(* Logix 5000 project; controller FV vendor 1 type 14 code 217 rev 31.11; software revision 31.00; part 32 of 63 *)
(* tags used below, declared in another part *)
   CWD : CHECKWORD_FLAGS;
   FR_data_file_value_to_move : DINT;
   FR_DEFOAM : PlantItem;   // DEFOAM
   FR_N120 : INT[265];   // YEAST CROP Yeast Cropping Main
   FR_N120_17_0_Storagebit : BOOL;
   FR_N120_17_1_Storagebit : BOOL;
   FR_N120_17_2_Storagebit : BOOL;
   FR_N120_17_3_Storagebit : BOOL;
   FR_N120_17_4_Storagebit : BOOL;
   FR_N120_17_5_Storagebit : BOOL;
   FR_N14 : INT[265];   // MVFV CIP Comms to MVFV CIP Un it PLC
   FR_N140 : INT[265];   // CIP
   FR_N150 : INT[265];   // Original N File From SLC, No Description Available
   FR_N20 : INT[265];   // GENERAL General Purpose Setp oints
   FR_N210 : INT[265];   // ANALOG_OUT Analog Outputs
   FR_N255 : INT[265];   // CHECKWORDS
   FR_N99 : INT[265];   // COMMENT Comment Lines
   FR_SFile : INT[255];   // SLC Equivalent System File, So Original Code Can Remain
   FR_T121 : TIMER[255];   // YEAST CROP
   FR_T144 : TIMER[255];   // CIP
   FR_T4 : TIMER[255];   // TIMER
   FR_VB1_AV02 : PlantItem;   // VB1_AV02
   FR_VB1_AV04 : PlantItem;   // VB1_AV04
   FR_VB1_AV07 : PlantItem;   // VB1_AV07
   FR_VB2_AV03 : PlantItem;   // VB2_AV03
   FR_VB3_AV03 : PlantItem;   // VB3_AV03
   FR_YC_1 : PlantItem;   // YC_1
   FR_YC_2 : PlantItem;   // YC_2
   FR_YC_IN2 : PlantItem;   // YC_IN2
   FR_YC_LL : PlantItem;   // YC_LL
   FR_YEAST_121_TEMPREAL : REAL;
   FR_YM_P01 : PlantItem;   // YM_P01
   FR_YM_P02 : PlantItem;   // YM_P02
   FR_YM_P03 : PlantItem;   // YM_P03
   FR_YP1_CIP : PlantItem;   // YP1_CIP
   FR_YP2_CIP : PlantItem;   // YP2_CIP
   FR_YP3_CIP : PlantItem;   // YP3_CIP
   scale_analog_result : REAL;
   Test_Cropping_done : BOOL;
(* FR_Common, continued *)

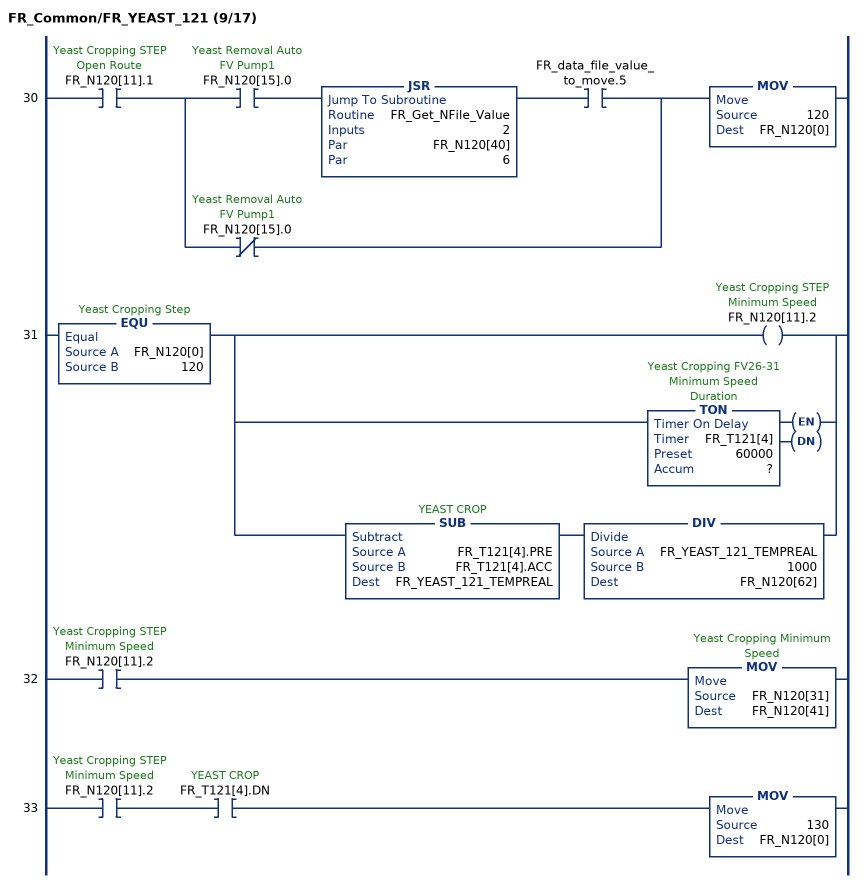
   30: XIC(FR_N120[11].1)[XIC(FR_N120[15].0) JSR(FR_Get_NFile_Value,2,FR_N120[40],6) XIC(FR_data_file_value_to_move.5) ,XIO(FR_N120[15].0) ]MOV(120,FR_N120[0]);
   31: EQU(FR_N120[0],120)[OTE(FR_N120[11].2) ,TON(FR_T121[4],?,?) ,SUB(FR_T121[4].PRE,FR_T121[4].ACC,FR_YEAST_121_TEMPREAL) DIV(FR_YEAST_121_TEMPREAL,1000,FR_N120[62]) ];
   32: XIC(FR_N120[11].2)MOV(FR_N120[31],FR_N120[41]);
   33: XIC(FR_N120[11].2)XIC(FR_T121[4].DN)MOV(130,FR_N120[0]);
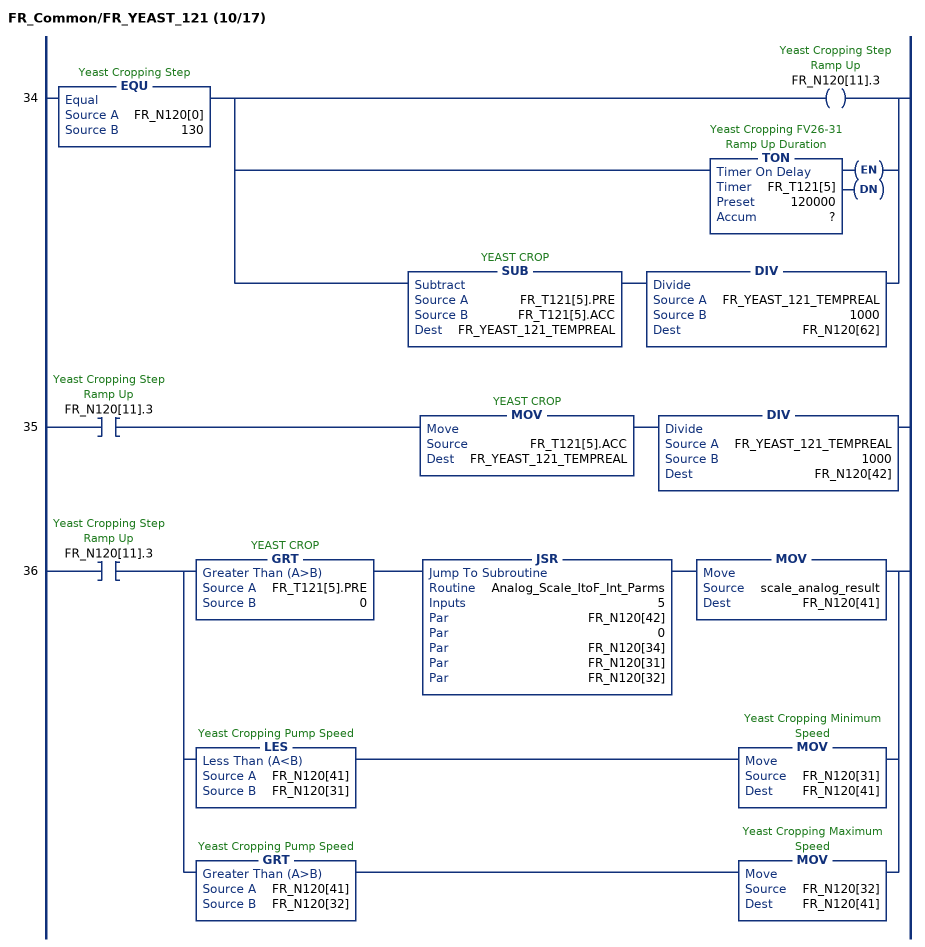
   34: EQU(FR_N120[0],130)[OTE(FR_N120[11].3) ,TON(FR_T121[5],?,?) ,SUB(FR_T121[5].PRE,FR_T121[5].ACC,FR_YEAST_121_TEMPREAL) DIV(FR_YEAST_121_TEMPREAL,1000,FR_N120[62]) ];
   35: XIC(FR_N120[11].3)MOV(FR_T121[5].ACC,FR_YEAST_121_TEMPREAL)DIV(FR_YEAST_121_TEMPREAL,1000,FR_N120[42]);
   36: XIC(FR_N120[11].3)[GRT(FR_T121[5].PRE,0) JSR(Analog_Scale_ItoF_Int_Parms,5,FR_N120[42],0,FR_N120[34],FR_N120[31],FR_N120[32]) MOV(scale_analog_result,FR_N120[41]) ,LES(FR_N120[41],FR_N120[31]) MOV(FR_N120[31],FR_N120[41]) ,GRT(FR_N120[41],FR_N120[32]) MOV(FR_N120[32],FR_N120[41]) ];
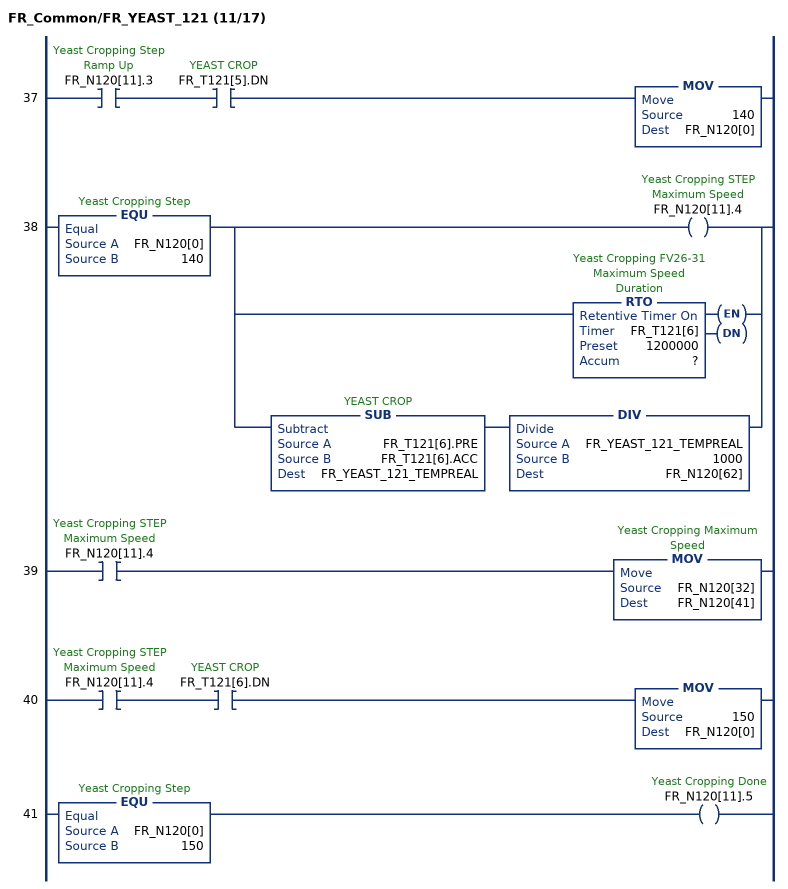
   37: XIC(FR_N120[11].3)XIC(FR_T121[5].DN)MOV(140,FR_N120[0]);
   38: EQU(FR_N120[0],140)[OTE(FR_N120[11].4) ,RTO(FR_T121[6],?,?) ,SUB(FR_T121[6].PRE,FR_T121[6].ACC,FR_YEAST_121_TEMPREAL) DIV(FR_YEAST_121_TEMPREAL,1000,FR_N120[62]) ];
   39: XIC(FR_N120[11].4)MOV(FR_N120[32],FR_N120[41]);
   40: XIC(FR_N120[11].4)XIC(FR_T121[6].DN)MOV(150,FR_N120[0]);
   41: EQU(FR_N120[0],150)OTE(FR_N120[11].5);
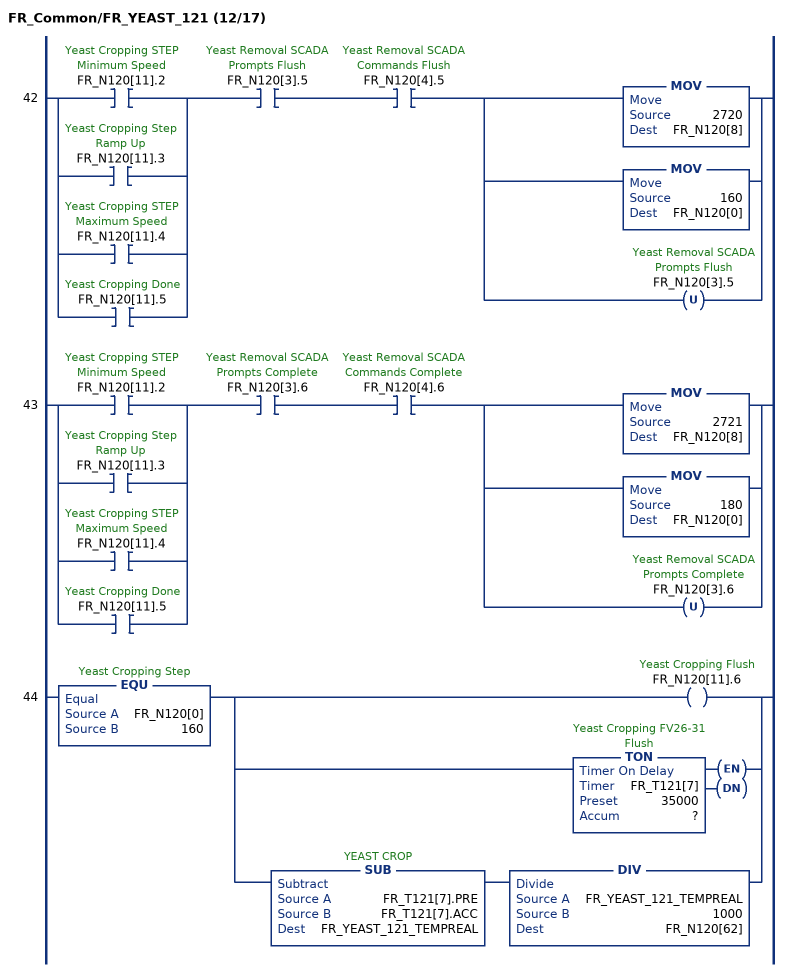
   42: [XIC(FR_N120[11].2) ,XIC(FR_N120[11].3) ,XIC(FR_N120[11].4) ,XIC(FR_N120[11].5) ]XIC(FR_N120[3].5)XIC(FR_N120[4].5)[MOV(2720,FR_N120[8]) ,MOV(160,FR_N120[0]) ,OTU(FR_N120[3].5) ];
   43: [XIC(FR_N120[11].2) ,XIC(FR_N120[11].3) ,XIC(FR_N120[11].4) ,XIC(FR_N120[11].5) ]XIC(FR_N120[3].6)XIC(FR_N120[4].6)[MOV(2721,FR_N120[8]) ,MOV(180,FR_N120[0]) ,OTU(FR_N120[3].6) ];
   44: EQU(FR_N120[0],160)[OTE(FR_N120[11].6) ,TON(FR_T121[7],?,?) ,SUB(FR_T121[7].PRE,FR_T121[7].ACC,FR_YEAST_121_TEMPREAL) DIV(FR_YEAST_121_TEMPREAL,1000,FR_N120[62]) ];
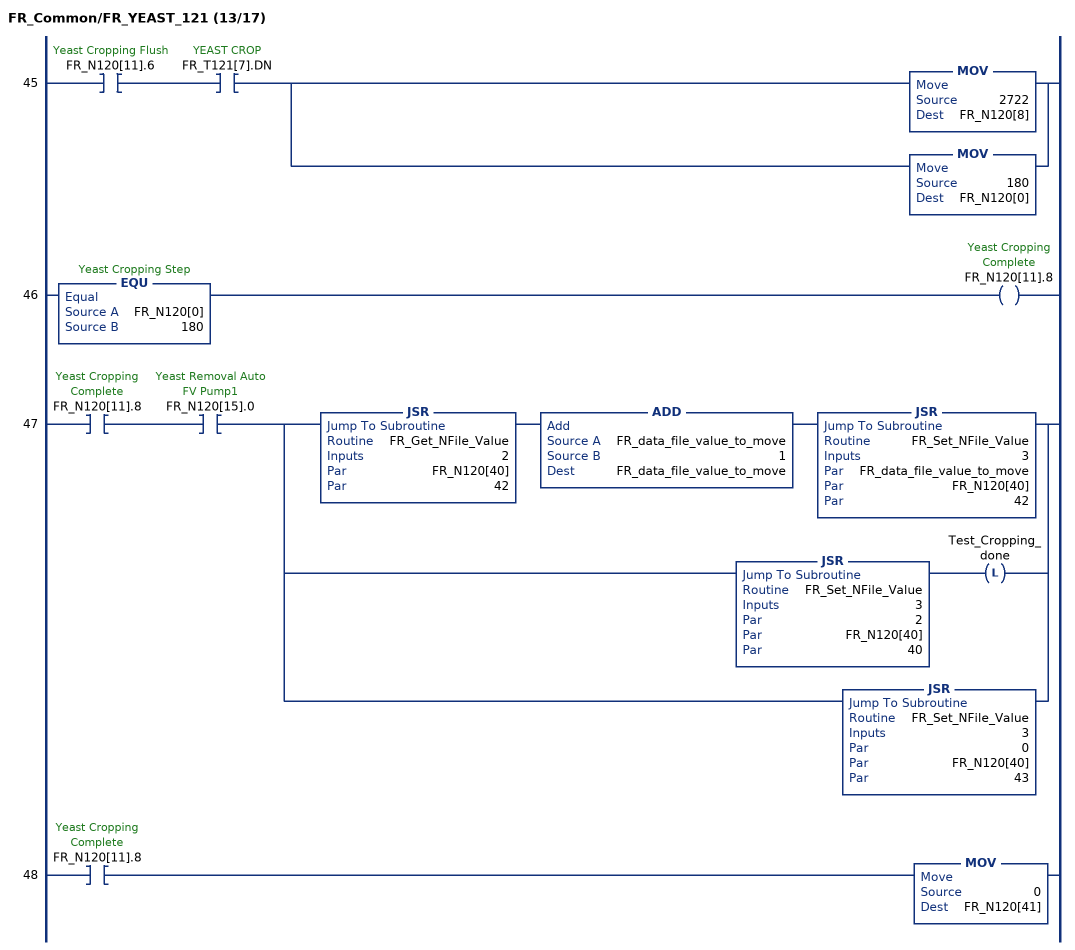
   45: XIC(FR_N120[11].6)XIC(FR_T121[7].DN)[MOV(2722,FR_N120[8]) ,MOV(180,FR_N120[0]) ];
   46: EQU(FR_N120[0],180)OTE(FR_N120[11].8);
   47: XIC(FR_N120[11].8)XIC(FR_N120[15].0)[JSR(FR_Get_NFile_Value,2,FR_N120[40],42) ADD(FR_data_file_value_to_move,1,FR_data_file_value_to_move) JSR(FR_Set_NFile_Value,3,FR_data_file_value_to_move,FR_N120[40],42) ,JSR(FR_Set_NFile_Value,3,2,FR_N120[40],40) OTL(Test_Cropping_done) ,JSR(FR_Set_NFile_Value,3,0,FR_N120[40],43) ];
   48: XIC(FR_N120[11].8)MOV(0,FR_N120[41]);
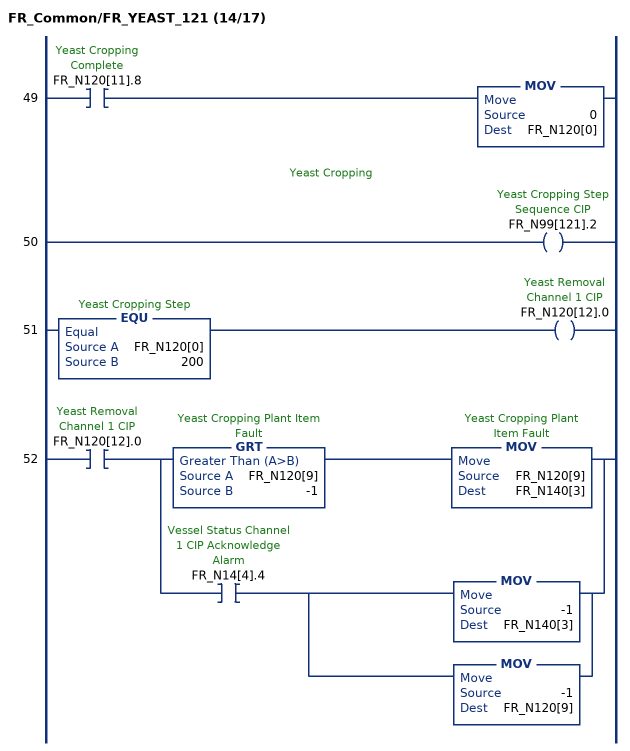
   49: XIC(FR_N120[11].8)MOV(0,FR_N120[0]);
   // Yeast Cropping
   50: OTE(FR_N99[121].2);
   51: EQU(FR_N120[0],200)OTE(FR_N120[12].0);
   52: XIC(FR_N120[12].0)[GRT(FR_N120[9],-1) MOV(FR_N120[9],FR_N140[3]) ,XIC(FR_N14[4].4) [MOV(-1,FR_N140[3]) ,MOV(-1,FR_N120[9]) ] ];
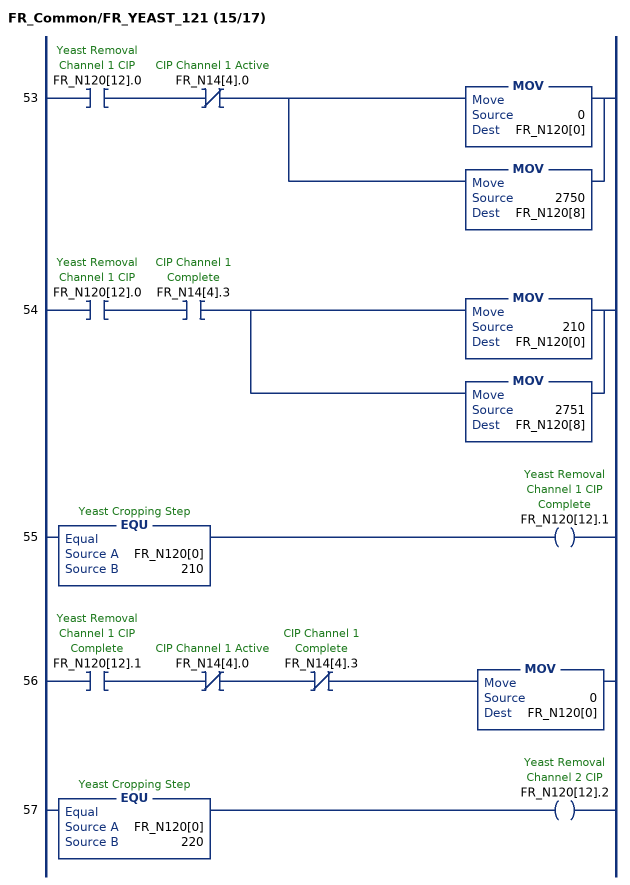
   53: XIC(FR_N120[12].0)XIO(FR_N14[4].0)[MOV(0,FR_N120[0]) ,MOV(2750,FR_N120[8]) ];
   54: XIC(FR_N120[12].0)XIC(FR_N14[4].3)[MOV(210,FR_N120[0]) ,MOV(2751,FR_N120[8]) ];
   55: EQU(FR_N120[0],210)OTE(FR_N120[12].1);
   56: XIC(FR_N120[12].1)XIO(FR_N14[4].0)XIO(FR_N14[4].3)MOV(0,FR_N120[0]);
   57: EQU(FR_N120[0],220)OTE(FR_N120[12].2);
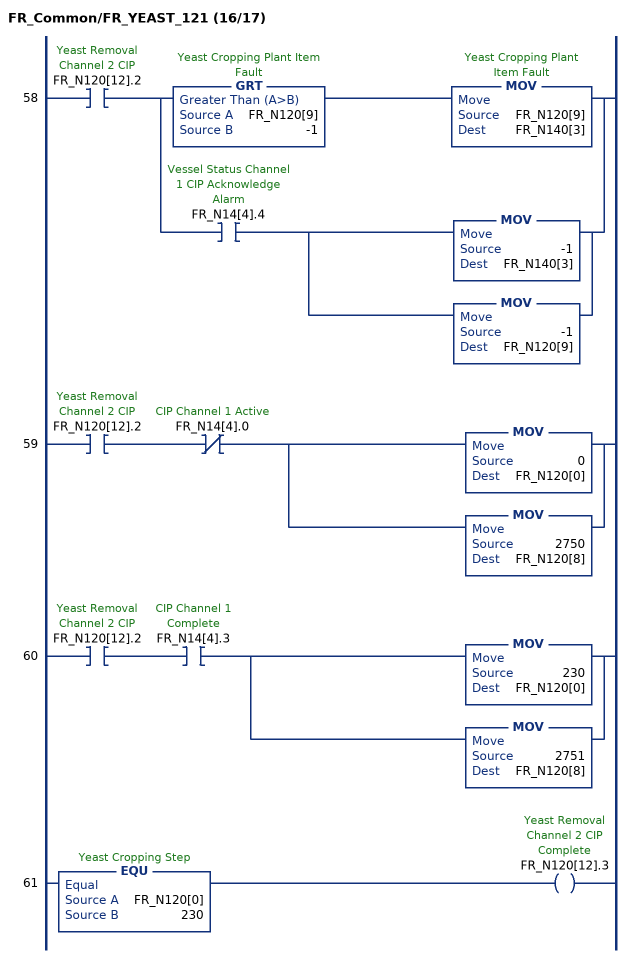
   58: XIC(FR_N120[12].2)[GRT(FR_N120[9],-1) MOV(FR_N120[9],FR_N140[3]) ,XIC(FR_N14[4].4) [MOV(-1,FR_N140[3]) ,MOV(-1,FR_N120[9]) ] ];
   59: XIC(FR_N120[12].2)XIO(FR_N14[4].0)[MOV(0,FR_N120[0]) ,MOV(2750,FR_N120[8]) ];
   60: XIC(FR_N120[12].2)XIC(FR_N14[4].3)[MOV(230,FR_N120[0]) ,MOV(2751,FR_N120[8]) ];
   61: EQU(FR_N120[0],230)OTE(FR_N120[12].3);
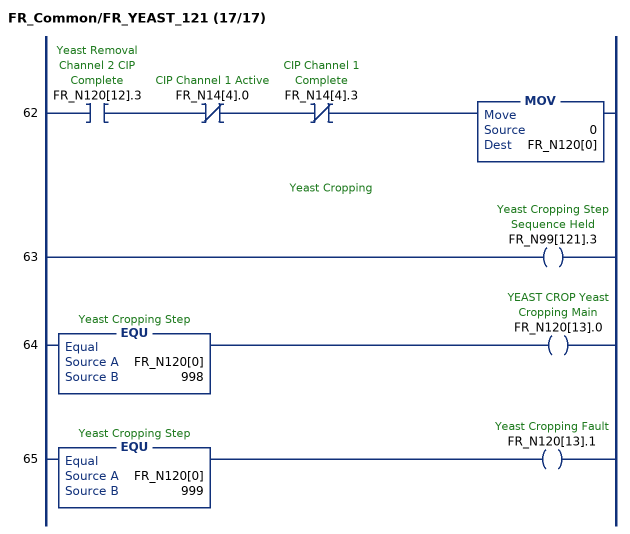
   62: XIC(FR_N120[12].3)XIO(FR_N14[4].0)XIO(FR_N14[4].3)MOV(0,FR_N120[0]);
   // Yeast Cropping
   63: OTE(FR_N99[121].3);
   64: EQU(FR_N120[0],998)OTE(FR_N120[13].0);
   65: EQU(FR_N120[0],999)OTE(FR_N120[13].1);
END_ROUTINE

ROUTINE FR_YEAST_COLL_150   (* ladder *)
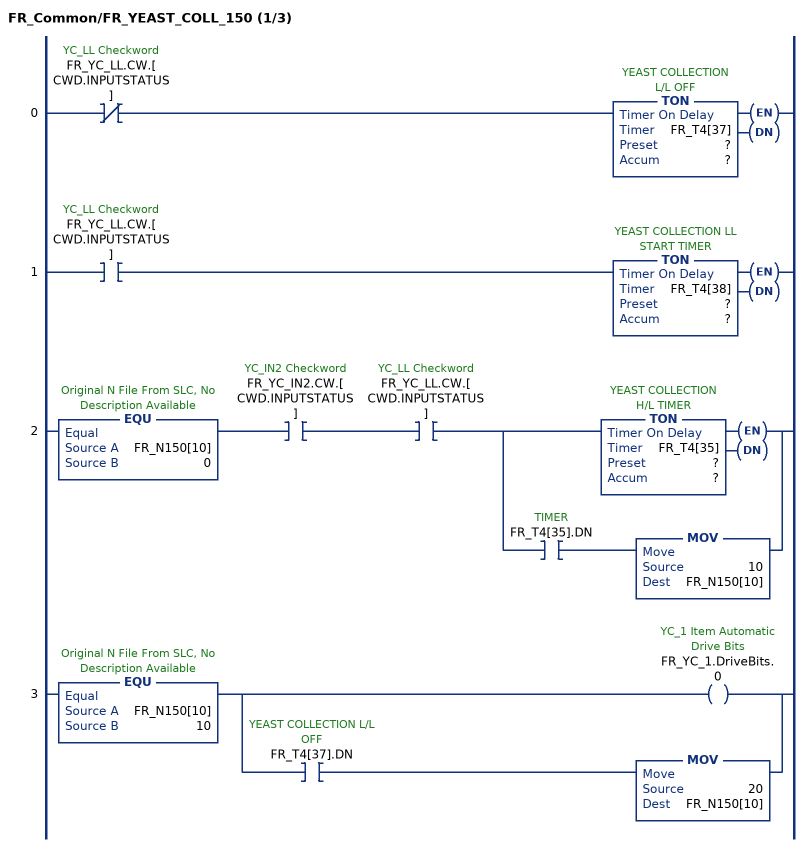
   0: XIO(FR_YC_LL.CW.[CWD.INPUTSTATUS])TON(FR_T4[37],?,?);
   1: XIC(FR_YC_LL.CW.[CWD.INPUTSTATUS])TON(FR_T4[38],?,?);
   2: EQU(FR_N150[10],0)XIC(FR_YC_IN2.CW.[CWD.INPUTSTATUS])XIC(FR_YC_LL.CW.[CWD.INPUTSTATUS])[TON(FR_T4[35],?,?) ,XIC(FR_T4[35].DN) MOV(10,FR_N150[10]) ];
   3: EQU(FR_N150[10],10)[OTE(FR_YC_1.DriveBits.0) ,XIC(FR_T4[37].DN) MOV(20,FR_N150[10]) ];
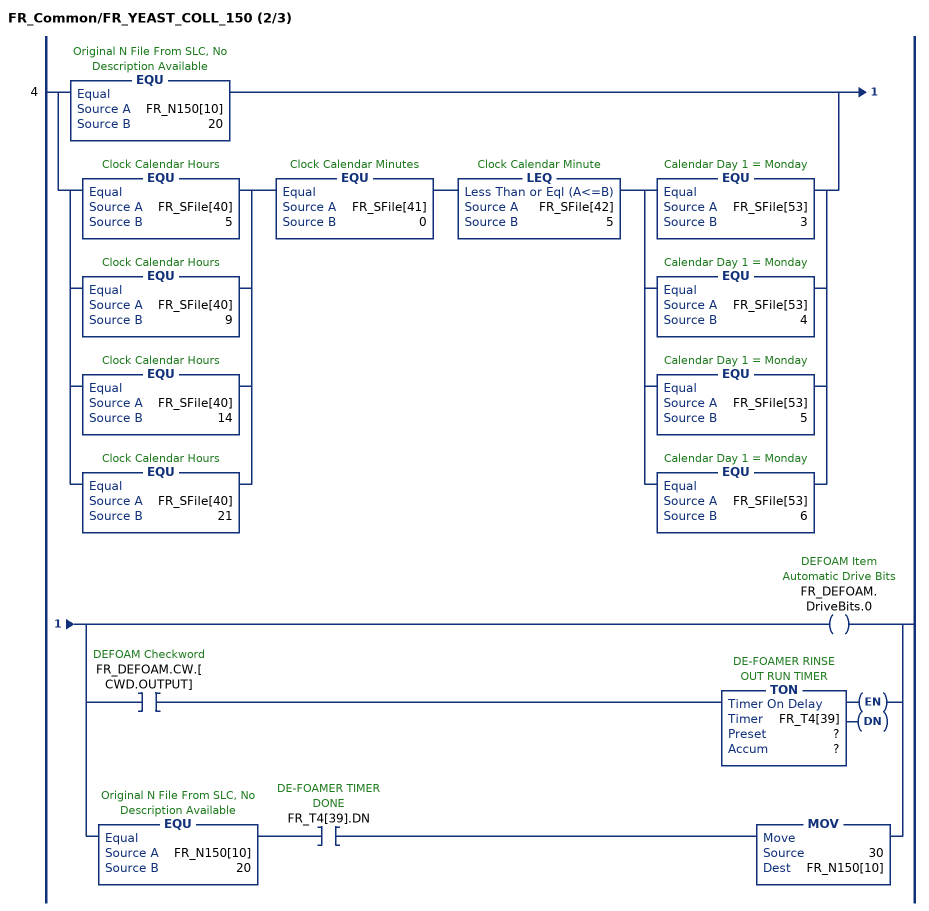
   4: [EQU(FR_N150[10],20) ,[EQU(FR_SFile[40],5) ,[EQU(FR_SFile[40],9) ,[EQU(FR_SFile[40],14) ,EQU(FR_SFile[40],21) ] ] ] EQU(FR_SFile[41],0) LEQ(FR_SFile[42],5) [EQU(FR_SFile[53],3) ,[EQU(FR_SFile[53],4) ,[EQU(FR_SFile[53],5) ,EQU(FR_SFile[53],6) ] ] ] ][OTE(FR_DEFOAM.DriveBits.0) ,[XIC(FR_DEFOAM.CW.[CWD.OUTPUT]) TON(FR_T4[39],?,?) ,EQU(FR_N150[10],20) XIC(FR_T4[39].DN) MOV(30,FR_N150[10]) ] ];
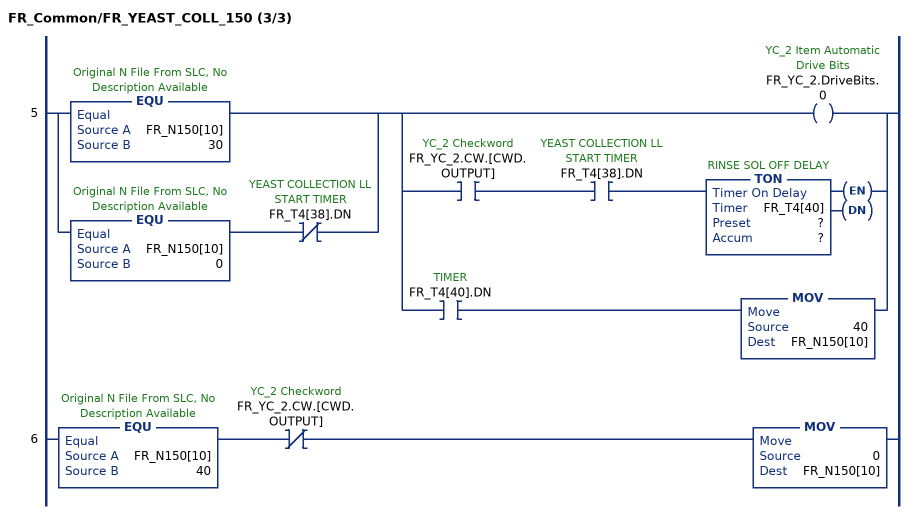
   5: [EQU(FR_N150[10],30) ,EQU(FR_N150[10],0) XIO(FR_T4[38].DN) ][OTE(FR_YC_2.DriveBits.0) ,[XIC(FR_YC_2.CW.[CWD.OUTPUT]) XIC(FR_T4[38].DN) TON(FR_T4[40],?,?) ,XIC(FR_T4[40].DN) MOV(40,FR_N150[10]) ] ];
   6: EQU(FR_N150[10],40)XIO(FR_YC_2.CW.[CWD.OUTPUT])MOV(0,FR_N150[10]);
END_ROUTINE

ROUTINE FR_YEAST_OP_122   (* ladder *)
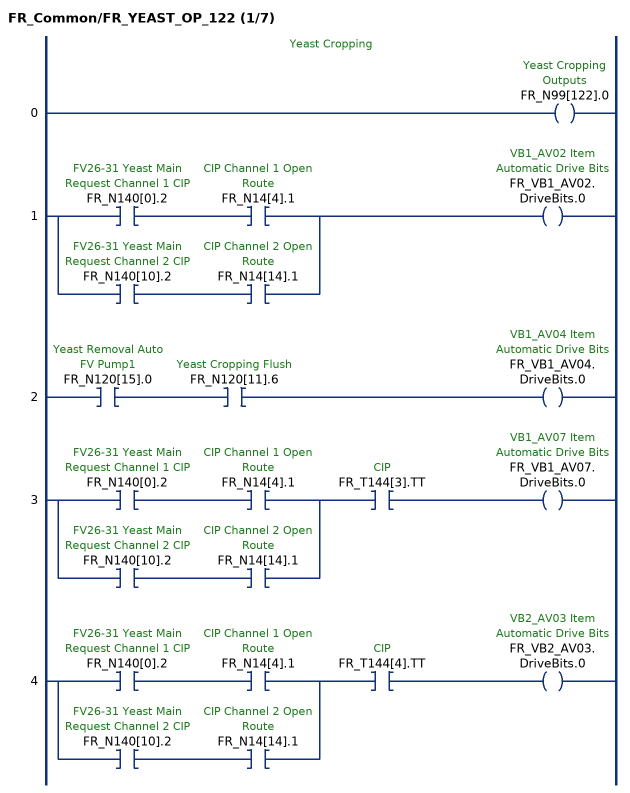
   // Yeast Cropping
   0: OTE(FR_N99[122].0);
   1: [XIC(FR_N140[0].2) XIC(FR_N14[4].1) ,XIC(FR_N140[10].2) XIC(FR_N14[14].1) ]OTE(FR_VB1_AV02.DriveBits.0);
   2: XIC(FR_N120[15].0)XIC(FR_N120[11].6)OTE(FR_VB1_AV04.DriveBits.0);
   3: [XIC(FR_N140[0].2) XIC(FR_N14[4].1) ,XIC(FR_N140[10].2) XIC(FR_N14[14].1) ]XIC(FR_T144[3].TT)OTE(FR_VB1_AV07.DriveBits.0);
   4: [XIC(FR_N140[0].2) XIC(FR_N14[4].1) ,XIC(FR_N140[10].2) XIC(FR_N14[14].1) ]XIC(FR_T144[4].TT)OTE(FR_VB2_AV03.DriveBits.0);
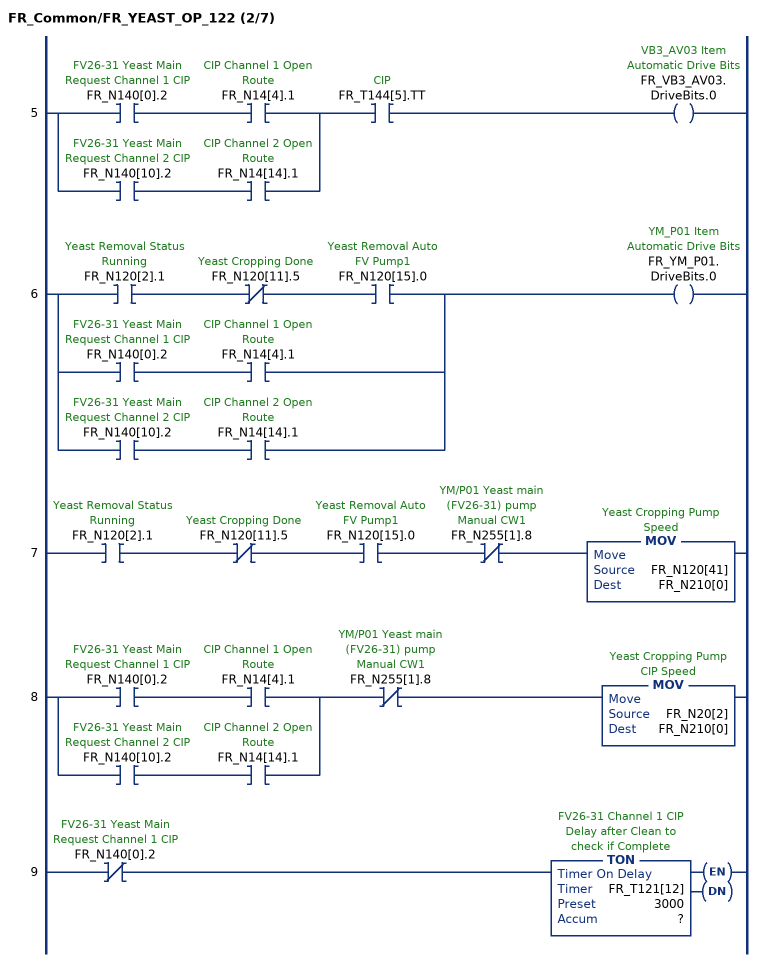
   5: [XIC(FR_N140[0].2) XIC(FR_N14[4].1) ,XIC(FR_N140[10].2) XIC(FR_N14[14].1) ]XIC(FR_T144[5].TT)OTE(FR_VB3_AV03.DriveBits.0);
   6: [XIC(FR_N120[2].1) XIO(FR_N120[11].5) XIC(FR_N120[15].0) ,XIC(FR_N140[0].2) XIC(FR_N14[4].1) ,XIC(FR_N140[10].2) XIC(FR_N14[14].1) ]OTE(FR_YM_P01.DriveBits.0);
   7: XIC(FR_N120[2].1)XIO(FR_N120[11].5)XIC(FR_N120[15].0)XIO(FR_N255[1].8)MOV(FR_N120[41],FR_N210[0]);
   8: [XIC(FR_N140[0].2) XIC(FR_N14[4].1) ,XIC(FR_N140[10].2) XIC(FR_N14[14].1) ]XIO(FR_N255[1].8)MOV(FR_N20[2],FR_N210[0]);
   9: XIO(FR_N140[0].2)TON(FR_T121[12],?,?);
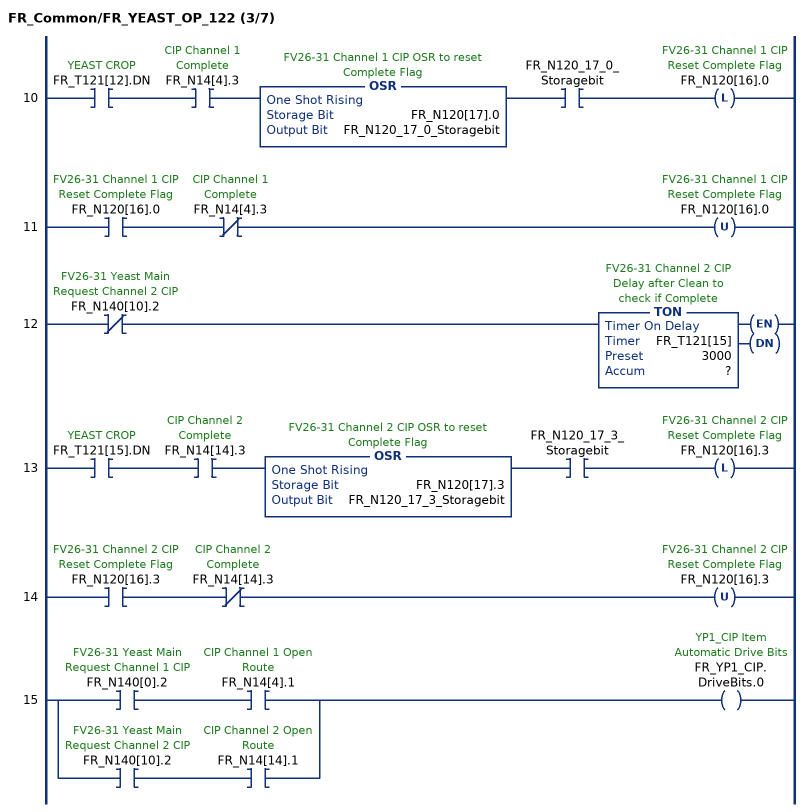
   10: XIC(FR_T121[12].DN)XIC(FR_N14[4].3)OSR(FR_N120[17].0,FR_N120_17_0_Storagebit)XIC(FR_N120_17_0_Storagebit)OTL(FR_N120[16].0);
   11: XIC(FR_N120[16].0)XIO(FR_N14[4].3)OTU(FR_N120[16].0);
   12: XIO(FR_N140[10].2)TON(FR_T121[15],?,?);
   13: XIC(FR_T121[15].DN)XIC(FR_N14[14].3)OSR(FR_N120[17].3,FR_N120_17_3_Storagebit)XIC(FR_N120_17_3_Storagebit)OTL(FR_N120[16].3);
   14: XIC(FR_N120[16].3)XIO(FR_N14[14].3)OTU(FR_N120[16].3);
   15: [XIC(FR_N140[0].2) XIC(FR_N14[4].1) ,XIC(FR_N140[10].2) XIC(FR_N14[14].1) ]OTE(FR_YP1_CIP.DriveBits.0);
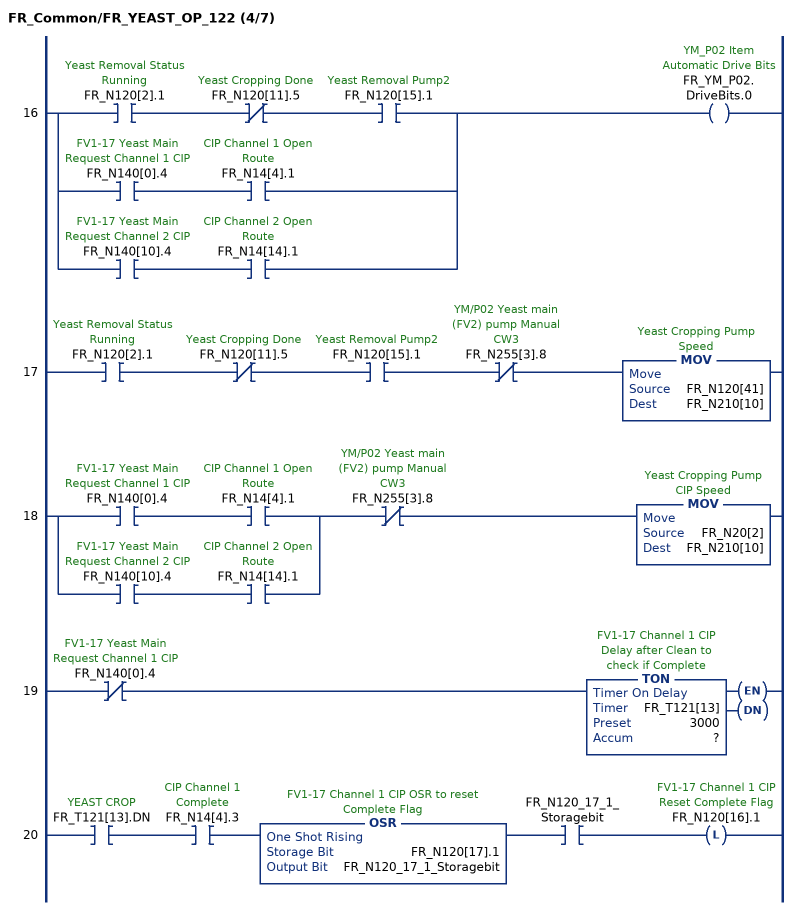
   16: [XIC(FR_N120[2].1) XIO(FR_N120[11].5) XIC(FR_N120[15].1) ,XIC(FR_N140[0].4) XIC(FR_N14[4].1) ,XIC(FR_N140[10].4) XIC(FR_N14[14].1) ]OTE(FR_YM_P02.DriveBits.0);
   17: XIC(FR_N120[2].1)XIO(FR_N120[11].5)XIC(FR_N120[15].1)XIO(FR_N255[3].8)MOV(FR_N120[41],FR_N210[10]);
   18: [XIC(FR_N140[0].4) XIC(FR_N14[4].1) ,XIC(FR_N140[10].4) XIC(FR_N14[14].1) ]XIO(FR_N255[3].8)MOV(FR_N20[2],FR_N210[10]);
   19: XIO(FR_N140[0].4)TON(FR_T121[13],?,?);
   20: XIC(FR_T121[13].DN)XIC(FR_N14[4].3)OSR(FR_N120[17].1,FR_N120_17_1_Storagebit)XIC(FR_N120_17_1_Storagebit)OTL(FR_N120[16].1);
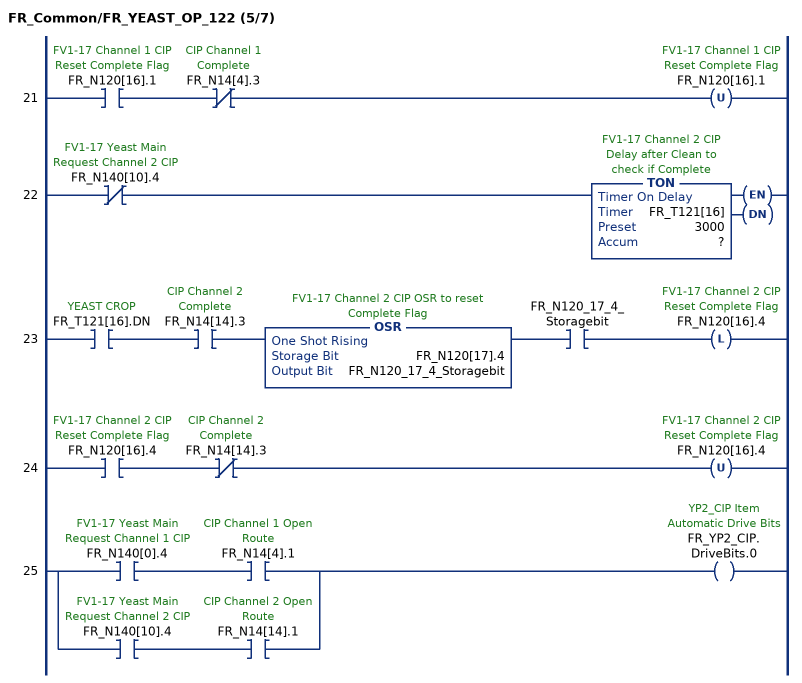
   21: XIC(FR_N120[16].1)XIO(FR_N14[4].3)OTU(FR_N120[16].1);
   22: XIO(FR_N140[10].4)TON(FR_T121[16],?,?);
   23: XIC(FR_T121[16].DN)XIC(FR_N14[14].3)OSR(FR_N120[17].4,FR_N120_17_4_Storagebit)XIC(FR_N120_17_4_Storagebit)OTL(FR_N120[16].4);
   24: XIC(FR_N120[16].4)XIO(FR_N14[14].3)OTU(FR_N120[16].4);
   25: [XIC(FR_N140[0].4) XIC(FR_N14[4].1) ,XIC(FR_N140[10].4) XIC(FR_N14[14].1) ]OTE(FR_YP2_CIP.DriveBits.0);
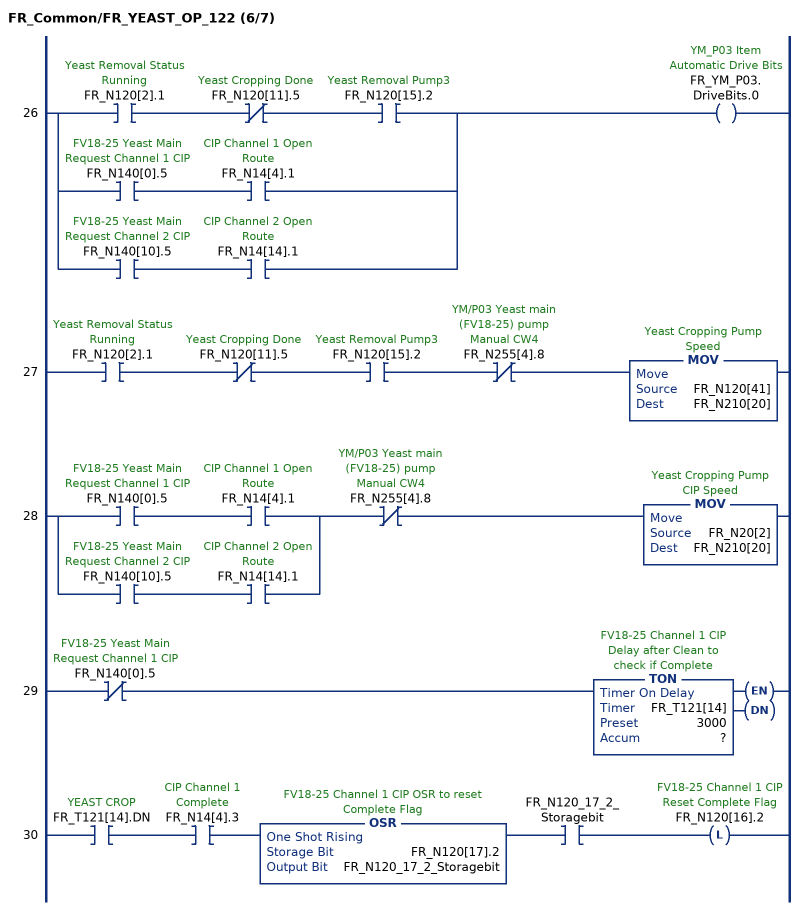
   26: [XIC(FR_N120[2].1) XIO(FR_N120[11].5) XIC(FR_N120[15].2) ,XIC(FR_N140[0].5) XIC(FR_N14[4].1) ,XIC(FR_N140[10].5) XIC(FR_N14[14].1) ]OTE(FR_YM_P03.DriveBits.0);
   27: XIC(FR_N120[2].1)XIO(FR_N120[11].5)XIC(FR_N120[15].2)XIO(FR_N255[4].8)MOV(FR_N120[41],FR_N210[20]);
   28: [XIC(FR_N140[0].5) XIC(FR_N14[4].1) ,XIC(FR_N140[10].5) XIC(FR_N14[14].1) ]XIO(FR_N255[4].8)MOV(FR_N20[2],FR_N210[20]);
   29: XIO(FR_N140[0].5)TON(FR_T121[14],?,?);
   30: XIC(FR_T121[14].DN)XIC(FR_N14[4].3)OSR(FR_N120[17].2,FR_N120_17_2_Storagebit)XIC(FR_N120_17_2_Storagebit)OTL(FR_N120[16].2);
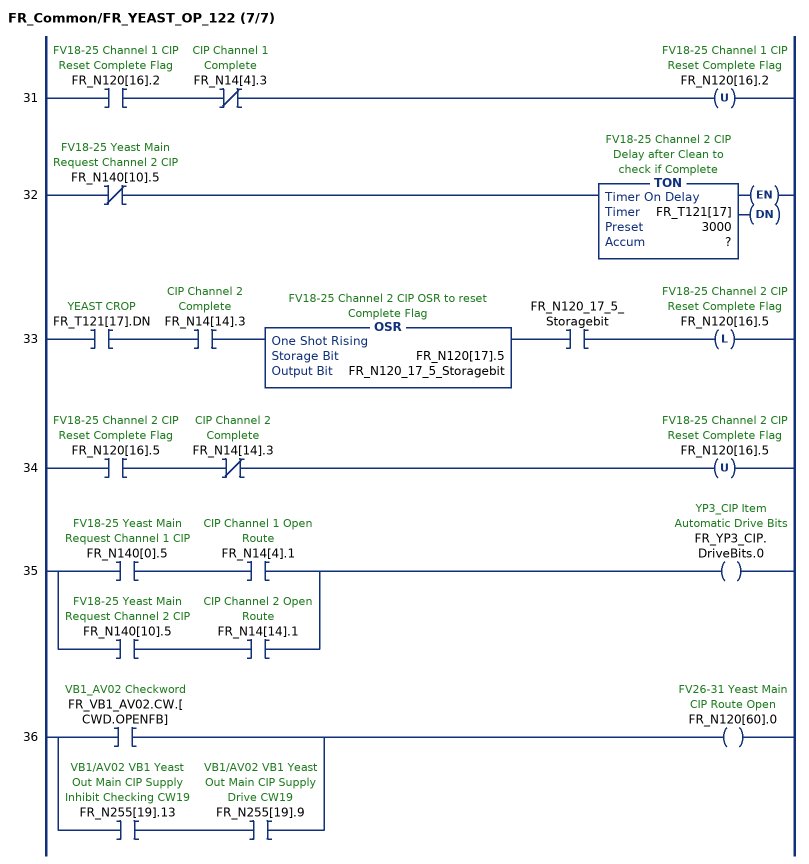
   31: XIC(FR_N120[16].2)XIO(FR_N14[4].3)OTU(FR_N120[16].2);
   32: XIO(FR_N140[10].5)TON(FR_T121[17],?,?);
   33: XIC(FR_T121[17].DN)XIC(FR_N14[14].3)OSR(FR_N120[17].5,FR_N120_17_5_Storagebit)XIC(FR_N120_17_5_Storagebit)OTL(FR_N120[16].5);
   34: XIC(FR_N120[16].5)XIO(FR_N14[14].3)OTU(FR_N120[16].5);
   35: [XIC(FR_N140[0].5) XIC(FR_N14[4].1) ,XIC(FR_N140[10].5) XIC(FR_N14[14].1) ]OTE(FR_YP3_CIP.DriveBits.0);
   36: [XIC(FR_VB1_AV02.CW.[CWD.OPENFB]) ,XIC(FR_N255[19].13) XIC(FR_N255[19].9) ]OTE(FR_N120[60].0);
END_ROUTINE
